(* Logix 5000 project; controller Seperator 1756-L85E rev 33.11; software revision 33.01 *)

TASK IO_Task (periodic, rate 250 ms, priority 2, watchdog 5000 ms) : IO_Simulation
TASK MainTask (continuous, watchdog 5000 ms) : Main_Sequencer, Filler, Capper, Capper_Heads, Filler_Heads1, Filler_Heads2, Filler_Heads3
TASK Process_Control (periodic, rate 250 ms, priority 2, watchdog 5000 ms) : Seperator_Control
TASK RandomTask (event, rate 1 ms, priority 1, watchdog 5000 ms) : RandomProgram   // Random Number Generator
TASK SignalGenerator (periodic, rate 100 ms, priority 1, watchdog 5000 ms) : RandomUpDown
TASK TemperatureLoops (periodic, rate 2000 ms, priority 3, watchdog 5000 ms) : TI101_Temperature

MODULES
   Local : 1756-L85E (ICP 0, rev 33.11)
END_MODULES

TYPE Benchmarks_Comparison :
STRUCT
   Actual_To_Baseline : REAL;
   Actual_To_Same_Interval_Prior_Periods : REAL;
   Production_Lines_To_Like_Lines : REAL;
   Production_Runs_To_Like_Runs : REAL;
END_STRUCT
END_TYPE

TYPE ControllerLEDStatus :
STRUCT
   Off : BOOL;
   SolidGreen : BOOL;
   FlashingGreen : BOOL;
   SolidYellow : BOOL;
   FlashingYellow : BOOL;
   FlashingRed : BOOL;
   SolidRed : BOOL;
END_STRUCT
END_TYPE

TYPE Facility :
STRUCT
   Company_Name : STRING;
   Location_Country : STRING;
   Location_State : STRING;
   Location_City : STRING;
   Benchmarks_Comparison : Benchmarks_Comparison;
   KPIs_Energy_PER_UOP : KPIs_Energy_PER_UOP;
   KPIs_GHG_PER_UOP : KPIs_GHG_PER_UOP;
   WAGES_Demand : WAGES_Demand;
   WAGES_Usage : WAGES_Usage;
END_STRUCT
END_TYPE

TYPE FaultRecord :
STRUCT
   timelow : DINT;
   timehigh : DINT;
   type : INT;
   code : INT;
   info : DINT[8];
END_STRUCT
END_TYPE

TYPE KPIs_Energy_PER_UOP :
STRUCT
   Eunits_PER_UOPunits : REAL;
   Edollar_PER_UOPunits : REAL;
   Eunits_PER_UOPdollar : REAL;
   Edollar_PER_UOPdollar : REAL;
END_STRUCT
END_TYPE

TYPE KPIs_GHG_PER_UOP :
STRUCT
   kG_CO2_e : REAL;
   Metric_Tonnes : REAL;
END_STRUCT
END_TYPE

TYPE Logix_Status_FP :
STRUCT
   ClearMinorFaults : DINT;
   Sts_MinorFaultEvents : DINT;
   Sts_MinorFaultBits : DINT;
   Sts_Redundant : DINT;
   Set_FaceplateAnimation : DINT;
   Val_ProductCode : DINT;
   MemoryTemp : INT[29];
   Val_raw_data : INT;
   Sts_IO_LED_raw : INT;
   Sts_ProductCode : INT;
   Val_Force_data_raw : INT;
   MemoryRequestData : SINT[12];
   Sts_Force_Installed : BOOL;
   Sts_Force_Enabled : BOOL;
   Sts_Faulted : BOOL;
   Sts_Run : BOOL;
   Sts_Program : BOOL;
   Sts_Minor_fault : BOOL;
   Sts_Major_fault : BOOL;
   Sts_KS_in_run : BOOL;
   Sts_KS_in_program : BOOL;
   Sts_KS_in_remote : BOOL;
   Sts_Changingmodes : BOOL;
   Sts_Test : BOOL;
   Sts_Ladder_Working : BOOL;
   Cmd_ClearFaultRecord : BOOL;
   Set_Controller_Description : STRING;
   UpdateDelayTimer : TIMER;
   Val_MajorFault : FaultRecord;
   Val_MFS : FaultRecord;
   Sts_IO_LED : ControllerLEDStatus;
   Sts_Battery_LED : ControllerLEDStatus;
   MemoryData : Memory_Data;
END_STRUCT
END_TYPE

TYPE Memory_Data :
STRUCT
   Free_Mem_IO : DINT;
   Free_Mem_DT : DINT;
   Free_Memory : DINT;
   Total_Mem_IO : DINT;
   Total_Mem_DT : DINT;
   Total_Memory : DINT;
   Biggest_IO_Mem_Size_Ava : DINT;
   Biggest_DT_Mem_Size_Ava : DINT;
END_STRUCT
END_TYPE

TYPE Motor :
STRUCT
   Start : BOOL;
   Stopped : BOOL;
   StartReq : BOOL;
   Alarm : BOOL;
   Running : BOOL;
END_STRUCT
END_TYPE

TYPE Moving_Analog_Indicator :
STRUCT
   Value : REAL;
   Medium_Alarm : REAL;
   High_Alarm : REAL;
   Min : REAL;
   Max : REAL;
END_STRUCT
END_TYPE

TYPE mtrcsdt :
STRUCT
   PartId : STRING;   // Static value per workcell
   IdealCT : REAL;   // Ideal time taken in Seconds to produce each Unit.
   GoodParts : DINT;   // Output Count in Units
   ScrapParts : DINT;   // Reject Count in Units
   TotalParts : DINT;   // Input Count in Units
   Running : BOOL;   // 1=Run Mode
   Monitored_Availability : BOOL;   // 1=Running OR Waiting
   Machine_State : INT;   // [0]=Undefined error [1]=Running [2]=Fault [3]=EfficiencyLoss
   BatchID : STRING;   // Product produced
   Colour : STRING;   // Product colour
   FaultEventTrigger : BOOL;   // 1=Fault detected
   FaultEventValue : INT;   // Fault code
   SlowEventTrigger : BOOL;   // 1=Workcell running slow
   SlowEventValue : INT;   // Slow reason code
   WarningEventTrigger : BOOL;   // 1=Warning detected
   WarningEventValue : INT;   // Warning code
END_STRUCT
END_TYPE

TYPE Phase_Control :
STRUCT
   Cmd_Start : BOOL;
   Cmd_Stop : BOOL;
   Cmd_Reset : BOOL;
END_STRUCT
END_TYPE

TYPE STRING_12 :
STRUCT
   LEN : DINT;
   DATA : SINT[12];
END_STRUCT
END_TYPE

TYPE STRING_16_UDT :
STRUCT
   LEN : DINT;
   DATA : SINT[16];
END_STRUCT
END_TYPE

TYPE STRING_20 :
STRUCT
   LEN : DINT;
   DATA : SINT[20];
END_STRUCT
END_TYPE

TYPE STRING_40 :
STRUCT
   LEN : DINT;
   DATA : SINT[40];
END_STRUCT
END_TYPE

TYPE Valve :
STRUCT
   Open : BOOL;
   Closed : BOOL;
   OpenReq : BOOL;
   Alarm : BOOL;
   Opened : BOOL;
END_STRUCT
END_TYPE

TYPE WAGES_Demand :
STRUCT
   Water_Demand : REAL;
   Air_Demand : REAL;
   Gas_Demand : REAL;
   Electric_Demand : REAL;
   Steam_Demand : REAL;
END_STRUCT
END_TYPE

TYPE WAGES_Usage :
STRUCT
   Water_Usage : REAL;
   Air_Usage : REAL;
   Gas_Usage : REAL;
   Electric_Usage : REAL;
   Steam_Usage : REAL;
END_STRUCT
END_TYPE

ADD_ON_INSTRUCTION AOI_SIM_RNG_Simple   (* revision 1.3, vendor Dr. Frank Jordan / Rockwell Automation, ExecutePrescan *)
// Simple Random Number Generator
// Revision note:
// This code is provided as application example without any warranty
// Help:
// George Marsaglia 's MWC (multiply with carry) algorithm
// (taken from http://www.codeproject.com/Articles/25172/Simple-Random-Number-Generation)
VAR_INPUT
   Seed : ALIAS FOR LocalSeed; {access Read Only, visible}
END_VAR
VAR_OUTPUT
   Count : DINT; {access Read Only, visible}
   Number : REAL; {access Read Only, visible}
END_VAR
VAR_INPUT
   TriggerSeed : ALIAS FOR LocalTriggerSeed; {access Read Only, visible}
   Reset : ALIAS FOR LocalReset; {access Read Only, visible}
END_VAR
VAR
   m_z : DINT; {access None}
   m_w : DINT; {access None}
   delta : REAL; {access None}
   consB : DINT; {access None}
   consA : DINT; {access None}
   AOI_UMUL : UMUL; {access None}
   u : DINT; {access None}
   AOI_UADD : UADD; {access None}
   LocalTriggerSeed : BOOL; {access Read Only}
   LocalSeed : DINT; {access Read Only}
   LocalReset : BOOL; {access Read Only}
   tmp : DINT; {access None}
   Overflow : BOOL; {access None}
END_VAR

ROUTINE Logic   (* ladder *)
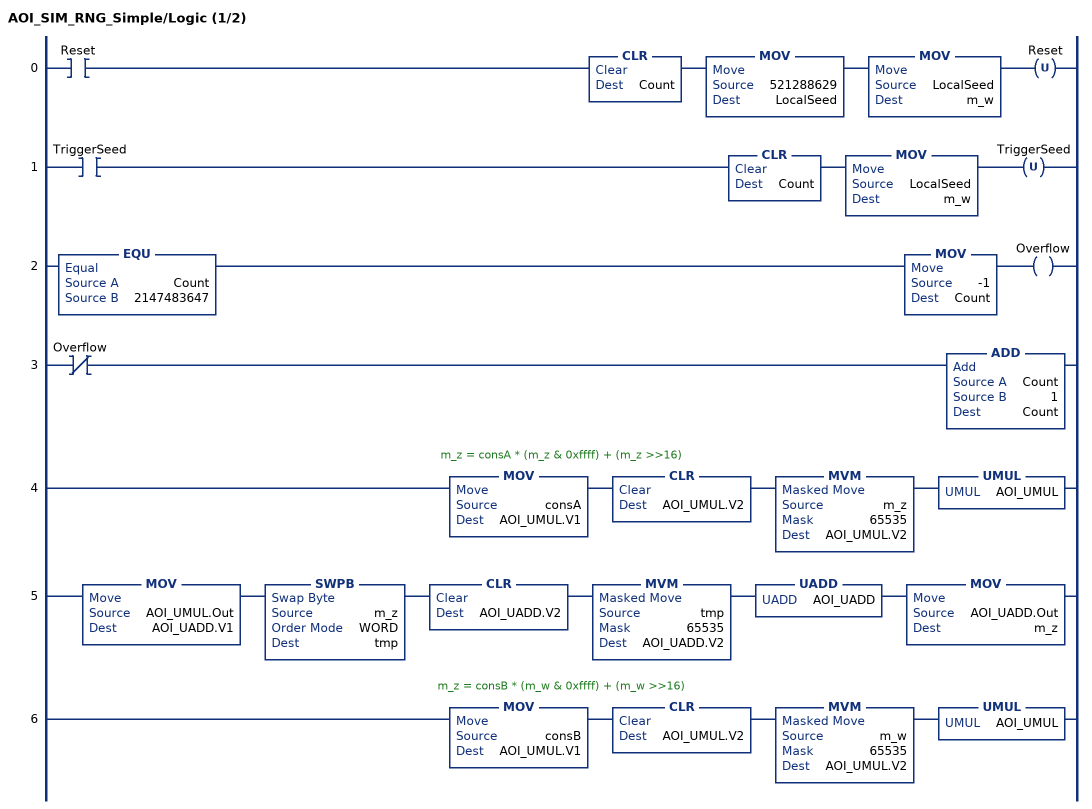
   0: XIC(Reset)CLR(Count)MOV(521288629,LocalSeed)MOV(LocalSeed,m_w)OTU(Reset);
   1: XIC(TriggerSeed)CLR(Count)MOV(LocalSeed,m_w)OTU(TriggerSeed);
   2: EQU(Count,2147483647)MOV(-1,Count)OTE(Overflow);
   3: XIO(Overflow)ADD(Count,1,Count);
   // m_z = consA * (m_z & 0xffff) + (m_z >>16)
   4: MOV(consA,AOI_UMUL.V1)CLR(AOI_UMUL.V2)MVM(m_z,65535,AOI_UMUL.V2)UMUL(AOI_UMUL);
   5: MOV(AOI_UMUL.Out,AOI_UADD.V1)SWPB(m_z,WORD,tmp)CLR(AOI_UADD.V2)MVM(tmp,65535,AOI_UADD.V2)UADD(AOI_UADD)MOV(AOI_UADD.Out,m_z);
   // m_z = consB * (m_w & 0xffff) + (m_w >>16)
   6: MOV(consB,AOI_UMUL.V1)CLR(AOI_UMUL.V2)MVM(m_w,65535,AOI_UMUL.V2)UMUL(AOI_UMUL);
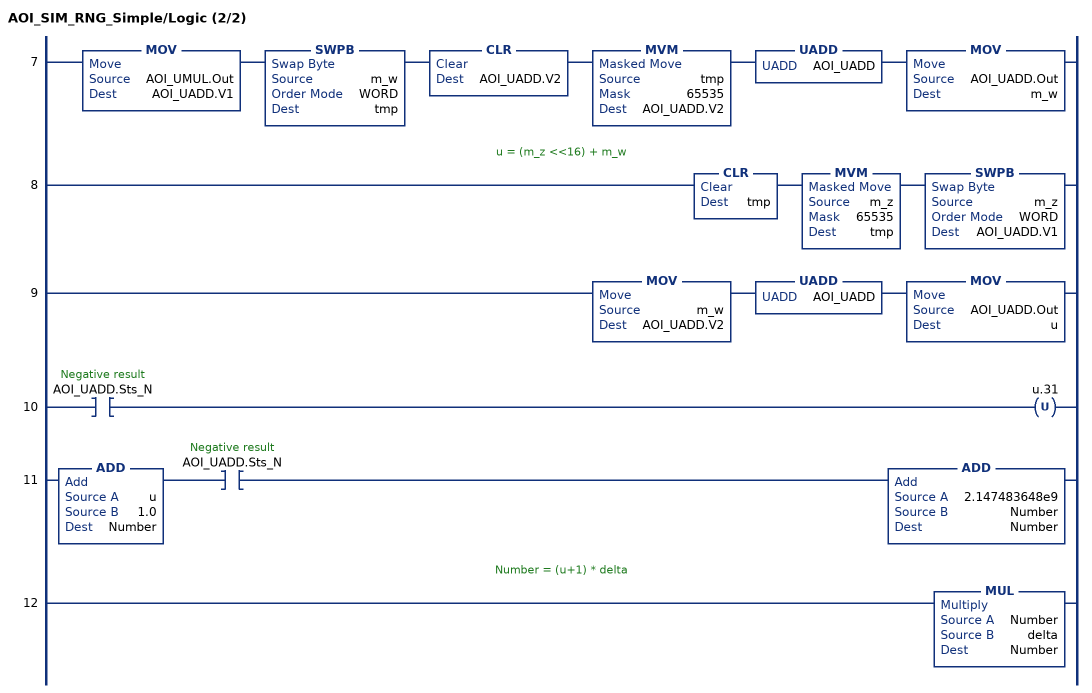
   7: MOV(AOI_UMUL.Out,AOI_UADD.V1)SWPB(m_w,WORD,tmp)CLR(AOI_UADD.V2)MVM(tmp,65535,AOI_UADD.V2)UADD(AOI_UADD)MOV(AOI_UADD.Out,m_w);
   // u = (m_z <<16) + m_w
   8: CLR(tmp)MVM(m_z,65535,tmp)SWPB(m_z,WORD,AOI_UADD.V1);
   9: MOV(m_w,AOI_UADD.V2)UADD(AOI_UADD)MOV(AOI_UADD.Out,u);
   10: XIC(AOI_UADD.Sts_N)OTU(u.31);
   11: ADD(u,1.0,Number)XIC(AOI_UADD.Sts_N)ADD(2.147483648e9,Number,Number);
   // Number = (u+1) * delta
   12: MUL(Number,delta,Number);
END_ROUTINE

ROUTINE Prescan   (* ladder *)
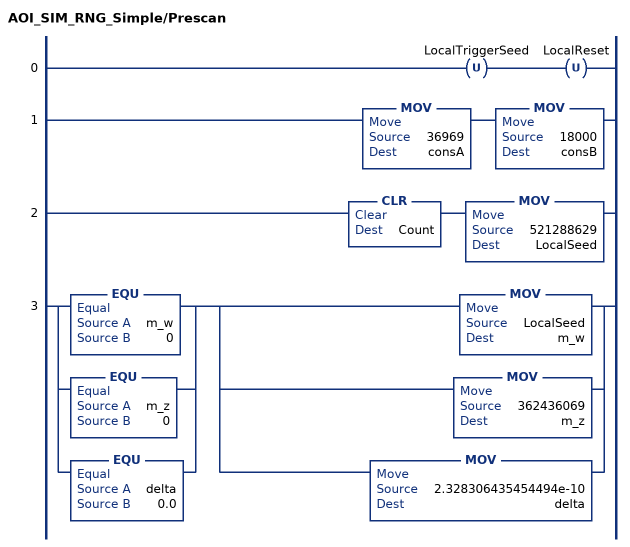
   0: OTU(LocalTriggerSeed)OTU(LocalReset);
   1: MOV(36969,consA)MOV(18000,consB);
   2: CLR(Count)MOV(521288629,LocalSeed);
   3: [EQU(m_w,0) ,EQU(m_z,0) ,EQU(delta,0.0) ][MOV(LocalSeed,m_w) ,MOV(362436069,m_z) ,MOV(2.328306435454494e-10,delta) ];
END_ROUTINE
END_ADD_ON_INSTRUCTION

ADD_ON_INSTRUCTION FTV_ctrl   (* revision 1.0 *)
VAR_INPUT
   nr_of_screens : DINT := 1; {visible}
   ActiveScreen : DINT;
   ScreenOverride : DINT;
   delay : DINT := 10; {visible}
   ScreenRequest : DINT;
END_VAR
VAR_OUTPUT
   Act : BOOL; {visible}
END_VAR
VAR
   Screen_delay : FBD_TIMER; {access None}
END_VAR

ROUTINE Logic   (* structured text *)
   Act:= (ActiveScreen >=100);
   
   Screen_delay.PRE:=delay*1000;
   Screen_delay.TimerEnable:=Act & NOT Screen_delay.DN & (ScreenRequest=0);
   TONR(Screen_delay);
   IF Act AND ScreenOverride<100 THEN ScreenOverride:=100;END_IF;
   IF Screen_delay.DN THEN ScreenOverride:= ScreenOverride+1;END_IF;
   IF ScreenOverride>=(100+ nr_of_screens) THEN ScreenOverride:=100;END_IF;
   
   IF ScreenRequest <> 0 THEN ScreenOverride:=ScreenRequest;
   	IF ActiveScreen=ScreenRequest THEN
   		ScreenOverride:=0;
   		ScreenRequest:=0;
   	END_IF;
   END_IF;
   
   IF NOT Act THEN ScreenOverride:=0; END_IF;
END_ROUTINE
END_ADD_ON_INSTRUCTION

ADD_ON_INSTRUCTION MotorSim   (* revision 1.0, vendor Rockwell, ExecutePrescan *)
VAR_INPUT
   MotorStartRequest : BOOL; {visible}
END_VAR
VAR_OUTPUT
   MotorRunning : BOOL; {access Read Only, visible}
   MotorStopped : BOOL; {access Read Only, visible}
END_VAR
VAR
   StartCommand : BOOL;
   RunningCommandDelay : TIMER := (PRE := 2000);
   StoppedCommandDelay : TIMER := (PRE := 2000);
END_VAR

ROUTINE Logic   (* ladder *)
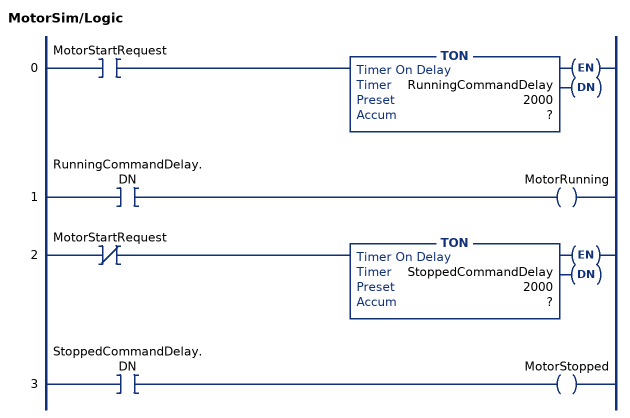
   0: XIC(MotorStartRequest)TON(RunningCommandDelay,?,?);
   1: XIC(RunningCommandDelay.DN)OTE(MotorRunning);
   2: XIO(MotorStartRequest)TON(StoppedCommandDelay,?,?);
   3: XIC(StoppedCommandDelay.DN)OTE(MotorStopped);
END_ROUTINE

ROUTINE Prescan   (* structured text *)
   RunningCommandDelay.PRE:=2000;
   StoppedCommandDelay.PRE:=2000;
   
END_ROUTINE
END_ADD_ON_INSTRUCTION

ADD_ON_INSTRUCTION P_Alarm   (* revision 3.0 02 Release, vendor Rockwell Automation, ExecutePrescan, ExecuteEnableInFalse *)
// Alarm
// Revision note:
// Changed suppress to shelve, inhibit to suppress (ISA 18.2-2009 and FTView 7 alignment), added auto unshelve timer, program command to unshelve. Removed: Ack on shelve. Added: clear Alm when disabled, PCfg_AllowExist, Cfg_Tag, Cfg_Cond, Inf_Lib, Inf_Type. Added Com_AE Local Tag for FTAE communication. Changed Cfg_MaxShelfT check to LEQ 0.  (INT 1 to 32767 is valid.)
// Help:
// Copyright © Rockwell Automation, Inc.  All Rights Reserved.
// This instruction monitors one input condition and provides one Alarm with:
//   * configurable latching (reset required) and acknowledgement requirement
//   * configurable alarm severity
//       1 = Low  (blue, typ. informational)
//       2 = Medium  (yelllow, typ. warning)
//       3 = High  (red, typ. process exception)
//       4 = Highest  (magenta, typ. equip. fault)
//   * configurable minimum ON time (e.g., to ensure it is seen by the HMI)
//   * commands to suppress/unsuppress (Prog), shelve/unshelve (Oper)
//         and disable/enable (Maint) the alarm.
//   * configurable amount of time shelved to automatically unshelve an alarm
//   * FTA&E support for suppressed, shelved and disabled states (V7.0)
// NOTE regarding parameter naming:
//   FTAE names (same as ALMD instruction) are used instead
//   of the ANSI/ISA 18.2-2009 names, as follows:
//    "Disabled" is the equivalent of "Out of Service" in ISA 18.2.
//       (The Disabled state is owned by Maintenance.)
//    "Suppressed" is the equivalent of "Suppressed by Design" in
//       ISA 18.2. (The Suppressed state is owned by Program logic.)
//    "Shelved" is the same as in ISA 18.2.
//       (The Shelved state is owned by Operator, but may be cleared
//       by Program logic based on time, shift change, etc.)
// This instruction is usually nested within other instructions, with one instance
// used for each Alarm generated by the containing instruction.  It may also be
// used as a standalone instruction for Alarm conditions generated by custom logic.
// FTAE Alarm Setup:
//   (object).(alarm).Com_AE.0:  Alarm to FTAE
//     .Com_AE.1:   Ack to/from FTAE
//     .Com_AE.3:   Shelved from FTAE Status
//     .Com_AE.4:   Shelve/Reshelve to FTAE Control (auto reset)
//     .Com_AE.5:   Unshelve to FTAE Control (auto reset)
//     .Com_AE.6:   Suppressed to/from FTAE
//     .Com_AE.8:   Unsuppress to FTAE Control (auto reset)
//     .Com_AE.9:   Disabled to/from FTAE
//     .Com_AE.11: Enable to FTAE Control (auto reset)
//    all other bits unused
//     .Cfg_MaxShelfT is also used in FTAE config.
VAR_INPUT
   Inp : BOOL := 1; {visible}   // Alarm Condition Input 1=Alarm
   Inp_Reset : BOOL; {visible}   // 1=Reset Alarm requiring reset
   Cfg_Exists : BOOL := 1;   // 1=Alarm configured to exist, 0=Does not exist, don't scan
   Cfg_ResetReqd : BOOL;   // 1=Latched Alarm, a Reset is required to clear this Alarm
   Cfg_AckReqd : BOOL := 1;   // 1=Acknowledge required for this Alarm
   Cfg_AllowShelve : BOOL := 1;   // 1=Allow Operator to Shelve this Alarm
   Cfg_AllowDisable : BOOL := 1;   // 1=Allow Maintenance to Disable this Alarm
   Cfg_PCmdClear : BOOL := 1;   // 1=Clear Program Commands on receipt 0=Leave Set
   Cfg_Severity : SINT := 3;   // Alarm Severity: 1=Low, 2=Medium, 3=High, 4=Highest
   Cfg_AlmMinOnT : DINT := 5;   // Minimum time Alm output stays on (sec)
   Cfg_MaxShelfT : INT := 480;   // Auto unshelve after shelved this long (1..32767 minutes)
   PCfg_AllowExist : BOOL := 1;   // 1=Alarm can be configured to exist, 0=other configs make alarm meaningless
   PCmd_Reset : BOOL;   // Program Command to Reset latched alarm
   PCmd_Ack : BOOL;   // Program Command to Acknowledge alarm
   PCmd_Suppress : BOOL;   // Program Command to Suppress by Design (inhibits new alarm)
   PCmd_Unsuppress : BOOL;   // Program Command to Unsuppress (allows new alarm)
   PCmd_Unshelve : BOOL;   // Program Command to Unshelve (e.g., on shift change)
   OCmd_Reset : BOOL;   // Operator Command to Reset latched alarm
   OCmd_Ack : BOOL;   // Operator Command to Acknowledge alarm
   OCmd_Shelve : BOOL;   // Operator Command to Shelve Alarm (inhibits new alarm)
   OCmd_Unshelve : BOOL;   // Operator Command to Unshelve alarm (allows new alarm)
   MCmd_Disable : BOOL;   // Maintenance Command to Disable alarm (inhibits new alarm)
   MCmd_Enable : BOOL;   // Maintenance Command to Enable alarm (allows new alarm)
END_VAR
VAR_OUTPUT
   Val_Notify : SINT; {access Read Only}   // Current Alarm Severity and Acknowledgement (enumeration)
   Val_MinToUnshelve : DINT; {access Read Only, visible}   // Number of minutes until this alarm unshelves itself (mmm:ss)
   Val_SecToUnshelve : DINT; {access Read Only, visible}   // Number of Seconds until this alarm unshelves itself (mmm:ss)
   Alm : ALIAS FOR Com_AE.0; {visible}   // Alarm output 1=In Alarm
   Ack : ALIAS FOR Com_AE.1; {visible}   // Alarm acknowledged status: 1=Ack rcvd
   Shelved : ALIAS FOR Com_AE.3; {visible}   // 1=Alarm has been Shelved by Operator (inhibits new alarm)
   Suppressed : ALIAS FOR Com_AE.6; {visible}   // 1=Alarm has been Suppressed by Program (inhibits new alarm)
   Disabled : ALIAS FOR Com_AE.9; {visible}   // 1=Alarm has been Disabled by Maintanance (inhibits new alarm)
   Sts_AlmInh : BOOL; {access Read Only}   // 1=Alarm has been suppressed, shelved or disabled, display "I" icon
   Sts_Err : BOOL; {access Read Only}   // 1=Error in Config: see detail Err_ bits for reason
   Err_Timer : BOOL; {access Read Only}   // 1=Error in Config: Alarm Min On Time, Shelf Time (use 0 to 2147483)
   Err_Severity : BOOL; {access Read Only}   // 1=Error in Config: Invalid Severity (use 1 to 4)
   Rdy_Reset : BOOL; {access Read Only}   // Ready to receive OCmd_Reset (enables button)
   Rdy_Ack : BOOL; {access Read Only}   // Ready to receive OCmd_Ack (enables button)
   Rdy_Shelve : BOOL; {access Read Only}   // Ready to receive OCmd_Shelve (enables button)
   Rdy_Unshelve : BOOL; {access Read Only}   // Ready to receive OCmd_Unshelve (enables button)
   Rdy_Disable : BOOL; {access Read Only}   // Ready to receive MCmd_Disable (enables button)
   Rdy_Enable : BOOL; {access Read Only}   // Ready to receive MCmd_Enable (enables button)
   P_Alarm : BOOL;   // Unique Parameter Name for auto - discovery
END_VAR
VAR
   Wrk_Alm : BOOL; {access None}   // Internal Alarm Status
   Wrk_Suppressed : BOOL; {access None}   // Internal Alarm Suppressed Status
   Wrk_AlmMinOnT : TIMER := (PRE := 5000); {access None}   // Alarm output minimum ON time to be seen by alarm server
   Wrk_AutoAckT : TIMER := (PRE := 5000); {access None}   // Time to clear Ack bit when Ack not required
   Wrk_ShelfT : TIMER; {access None}   // Time to auto Unshelve a Shelved Alarm
   Inf_Tab : SINT;   // Tab to display (FTView ME)
   Com_AE : INT := 2#0000_0000_0000_0010;   // Communication with HMI / Alarm/Event Server (see bit descriptions)
        .10   // (not used)
        .11   // Enable to AE Control
        .12   // (not used)
        .13   // (not used)
        .14   // (not used)
        .15   // (not used)
        .0   // Alarm to AE
        .1   // Acked from AE Status, Ack to AE Control
        .2   // (not used)
        .3   // Shelved from AE Status
        .4   // Shelve to AE Control
        .5   // Unshelve to AE Control
        .6   // Suppressed from AE Status, Suppress to AE Control
        .7   // (not used)
        .8   // Unsuppress to AE Control
        .9   // Disabled from AE Status, Disable to AE Control
   Cfg_Tag : STRING_20 := 'P_Alarm';   // Alarm Tag Text (e.g., "LAHH-101")
   Cfg_Cond : STRING_20 := 'Alarm Condition';   // Alarm Condition Text (e.g., "High-High PV")
   Wrk_SecToUnshelve : DINT; {access None}   // Number of seconds until this alarm unshelves itself
   Inf_Lib : STRING_12 := 'RA-BAS'; {access Read Only}   // Display Library for Faceplate call-up
   Inf_Type : STRING_16_UDT := 'P_Alarm'; {access Read Only}   // Must contain AOI name, used for HMI and Information S/W
END_VAR

ROUTINE EnableInFalse   (* ladder *)
// Perform Alarm processing, but Invert Alarm Input ("Inp") for use on LD rung (EnableIn False)
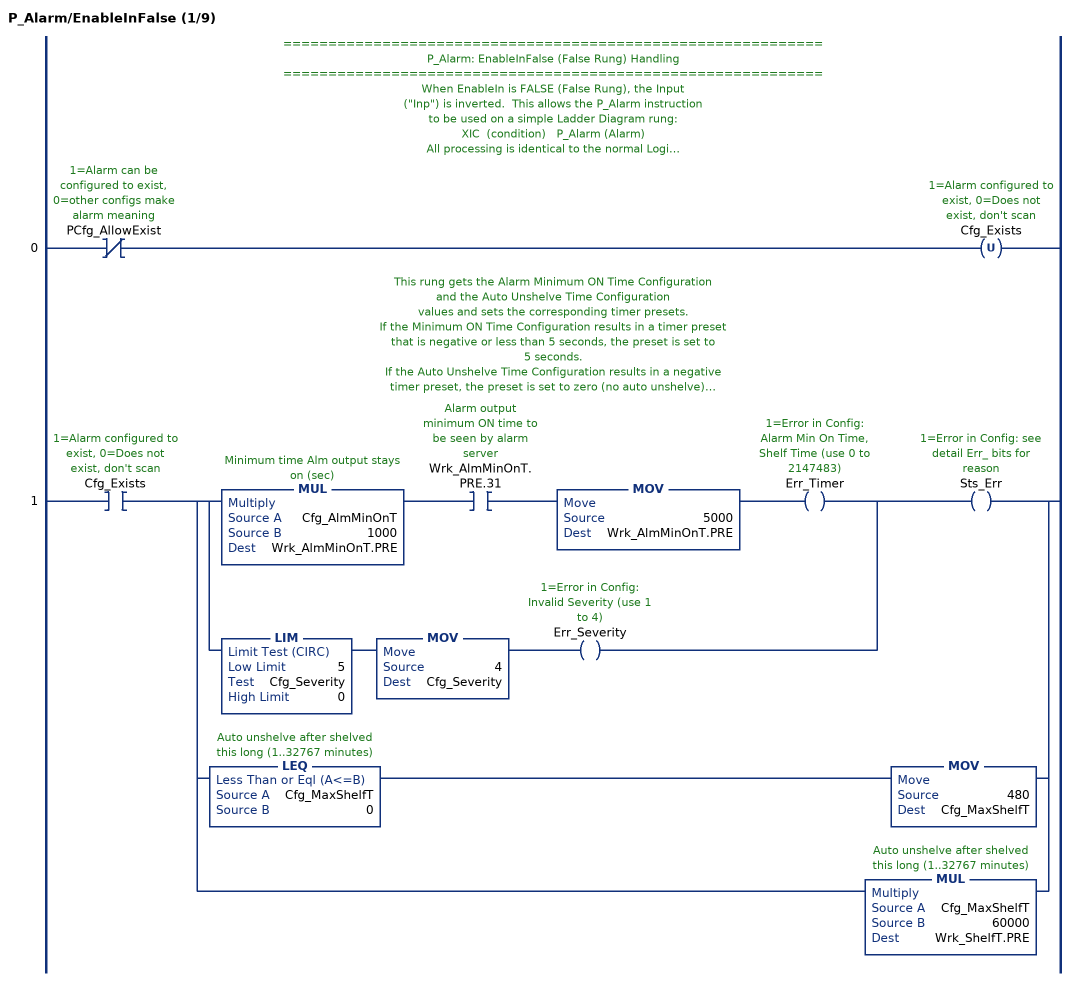
   // ============================================================
   // P_Alarm: EnableInFalse (False Rung) Handling
   // ============================================================
   // When EnableIn is FALSE (False Rung), the Input
   // ("Inp") is inverted.  This allows the P_Alarm instruction
   // to be used on a simple Ladder Diagram rung:
   // XIC  (condition)   P_Alarm (Alarm)
   // All processing is identical to the normal Logic
   // routine, except references to Inp are inverted!
   // ============================================================
   // CONFIGURATION
   // ============================================================
   // In the object containing this alarm, other configuration (such as not having
   // any limit switches) may make this particular alarm meaningless.
   // The Program Configuration "Allow Exist" is used to hide this alarm
   // on the object's faceplate and other graphics, and forces the Cfg_Exist to 0.
   // #####  V3.0-00  2013-06-30:  Added PCfg_AllowExist.  #####
   0: XIO(PCfg_AllowExist)OTU(Cfg_Exists);
   // This rung gets the Alarm Minimum ON Time Configuration
   // and the Auto Unshelve Time Configuration
   // values and sets the corresponding timer presets.
   // If the Minimum ON Time Configuration results in a timer preset
   // that is negative or less than 5 seconds, the preset is set to
   // 5 seconds.
   // If the Auto Unshelve Time Configuration results in a negative
   // timer preset, the preset is set to zero (no auto unshelve).
   //   The bad Config is flagged (Err_Timer).
   // Bad Config is also flagged if the Cfg_Severity is out of range (valid = 1..4)
   // #####  V3.0-00  2013-06-30:  Changed Program Inhibit to Suppress, Operator Suppress to Shelve.  #####
   // #####  Added Shelf Timer config check; if Severity out of range, make it "Fault".  #####
   // #####  V3.0-02  2013-10-30:  Changed Cfg_MaxShelfT check to LEQ 0.  (INT 1 to 32767 is valid.)  #####
   1: XIC(Cfg_Exists)[[MUL(Cfg_AlmMinOnT,1000,Wrk_AlmMinOnT.PRE) XIC(Wrk_AlmMinOnT.PRE.31) MOV(5000,Wrk_AlmMinOnT.PRE) OTE(Err_Timer) ,LIM(5,Cfg_Severity,0) MOV(4,Cfg_Severity) OTE(Err_Severity) ] OTE(Sts_Err) ,LEQ(Cfg_MaxShelfT,0) MOV(480,Cfg_MaxShelfT) ,MUL(Cfg_MaxShelfT,60000,Wrk_ShelfT.PRE) ];
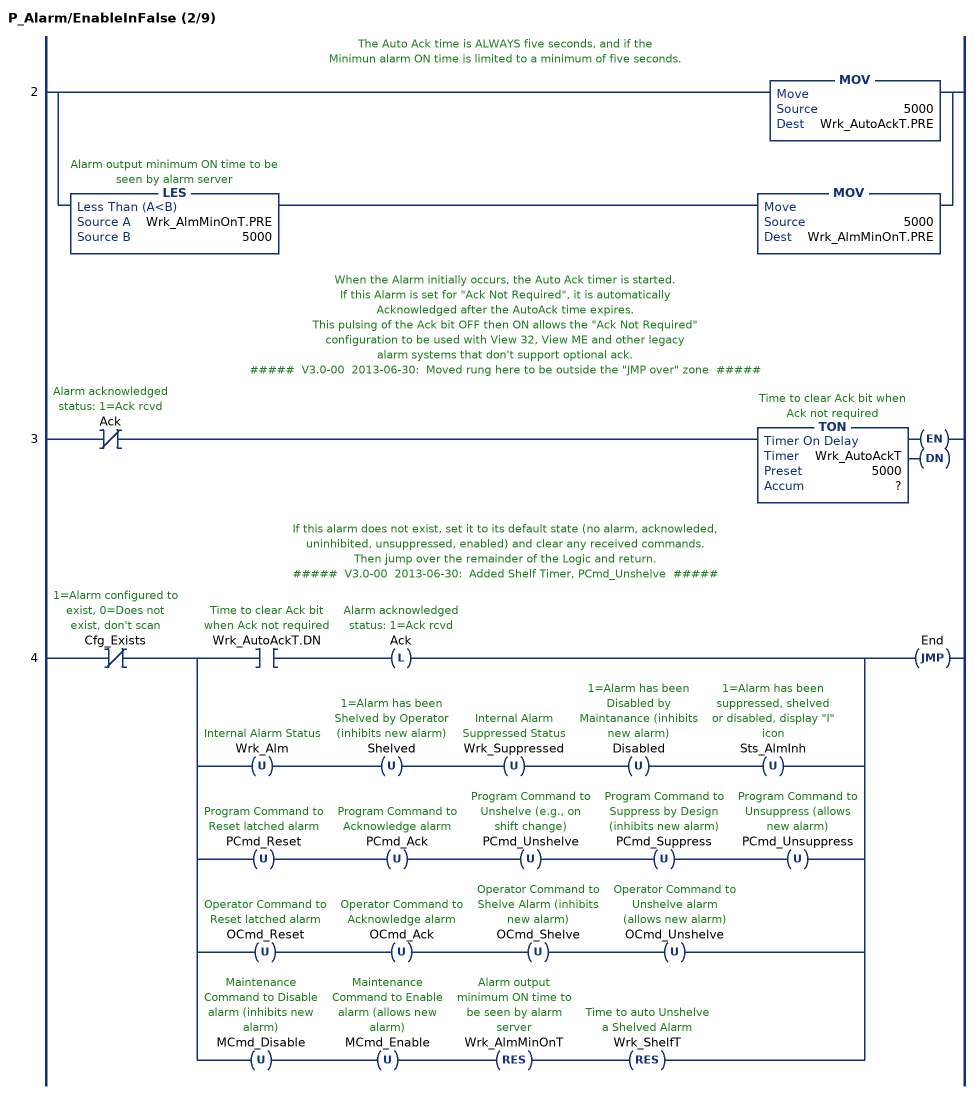
   // The Auto Ack time is ALWAYS five seconds, and if the
   // Minimun alarm ON time is limited to a minimum of five seconds.
   2: [MOV(5000,Wrk_AutoAckT.PRE) ,LES(Wrk_AlmMinOnT.PRE,5000) MOV(5000,Wrk_AlmMinOnT.PRE) ];
   // When the Alarm initially occurs, the Auto Ack timer is started.
   // If this Alarm is set for "Ack Not Required", it is automatically
   // Acknowledged after the AutoAck time expires.
   // This pulsing of the Ack bit OFF then ON allows the "Ack Not Required"
   // configuration to be used with View 32, View ME and other legacy
   // alarm systems that don't support optional ack.
   // #####  V3.0-00  2013-06-30:  Moved rung here to be outside the "JMP over" zone  #####
   3: XIO(Ack)TON(Wrk_AutoAckT,?,?);
   // If this alarm does not exist, set it to its default state (no alarm, acknowleded,
   // uninhibited, unsuppressed, enabled) and clear any received commands.
   // Then jump over the remainder of the Logic and return.
   // #####  V3.0-00  2013-06-30:  Added Shelf Timer, PCmd_Unshelve  #####
   4: XIO(Cfg_Exists)[XIC(Wrk_AutoAckT.DN) OTL(Ack) ,OTU(Wrk_Alm) OTU(Shelved) OTU(Wrk_Suppressed) OTU(Disabled) OTU(Sts_AlmInh) ,OTU(PCmd_Reset) OTU(PCmd_Ack) OTU(PCmd_Unshelve) OTU(PCmd_Suppress) OTU(PCmd_Unsuppress) ,OTU(OCmd_Reset) OTU(OCmd_Ack) OTU(OCmd_Shelve) OTU(OCmd_Unshelve) ,OTU(MCmd_Disable) OTU(MCmd_Enable) RES(Wrk_AlmMinOnT) RES(Wrk_ShelfT) ]JMP(End);
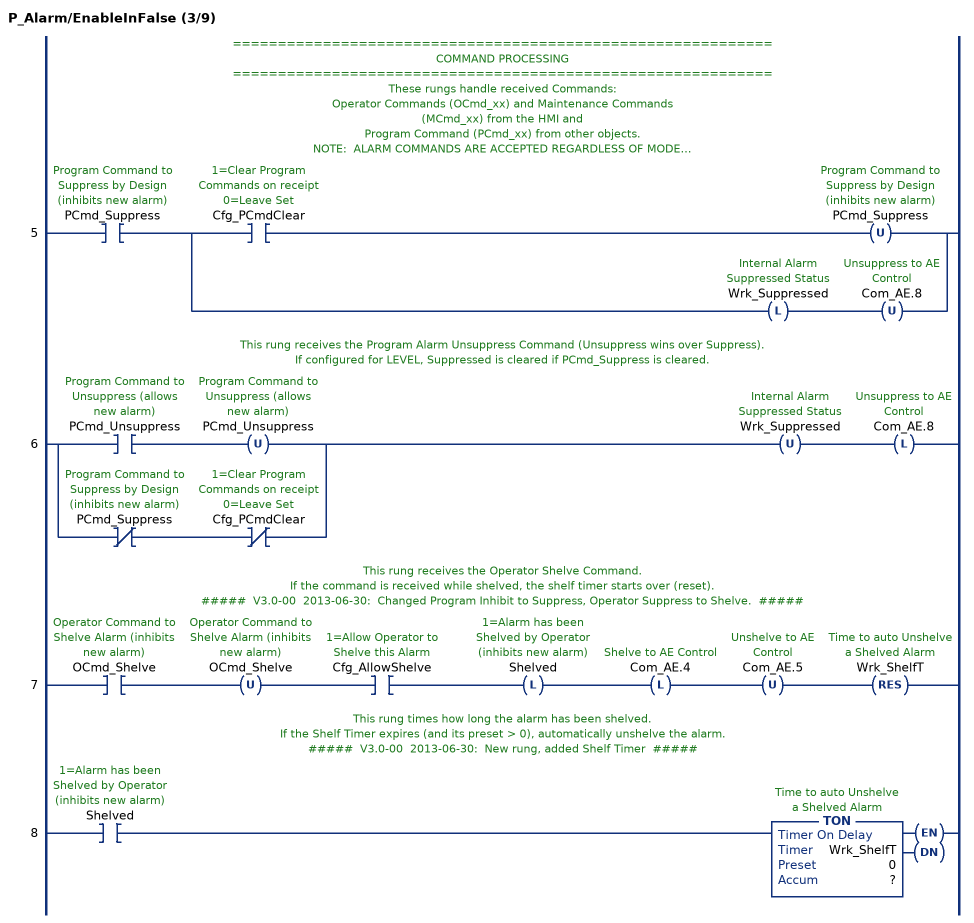
   // ============================================================
   // COMMAND PROCESSING
   // ============================================================
   // These rungs handle received Commands:
   // Operator Commands (OCmd_xx) and Maintenance Commands
   // (MCmd_xx) from the HMI and
   // Program Command (PCmd_xx) from other objects.
   // NOTE:  ALARM COMMANDS ARE ACCEPTED REGARDLESS OF MODE.
   // This rung receives the Program Alarm Inhibit Command.
   // If configured for EDGE, the Command is cleared.
   5: XIC(PCmd_Suppress)[XIC(Cfg_PCmdClear) OTU(PCmd_Suppress) ,OTL(Wrk_Suppressed) OTU(Com_AE.8) ];
   // This rung receives the Program Alarm Unsuppress Command (Unsuppress wins over Suppress).
   // If configured for LEVEL, Suppressed is cleared if PCmd_Suppress is cleared.
   6: [XIC(PCmd_Unsuppress) OTU(PCmd_Unsuppress) ,XIO(PCmd_Suppress) XIO(Cfg_PCmdClear) ]OTU(Wrk_Suppressed)OTL(Com_AE.8);
   // This rung receives the Operator Shelve Command.
   // If the command is received while shelved, the shelf timer starts over (reset).
   // #####  V3.0-00  2013-06-30:  Changed Program Inhibit to Suppress, Operator Suppress to Shelve.  #####
   7: XIC(OCmd_Shelve)OTU(OCmd_Shelve)XIC(Cfg_AllowShelve)OTL(Shelved)OTL(Com_AE.4)OTU(Com_AE.5)RES(Wrk_ShelfT);
   // This rung times how long the alarm has been shelved.
   // If the Shelf Timer expires (and its preset > 0), automatically unshelve the alarm.
   // #####  V3.0-00  2013-06-30:  New rung, added Shelf Timer  #####
   8: XIC(Shelved)TON(Wrk_ShelfT,?,?);
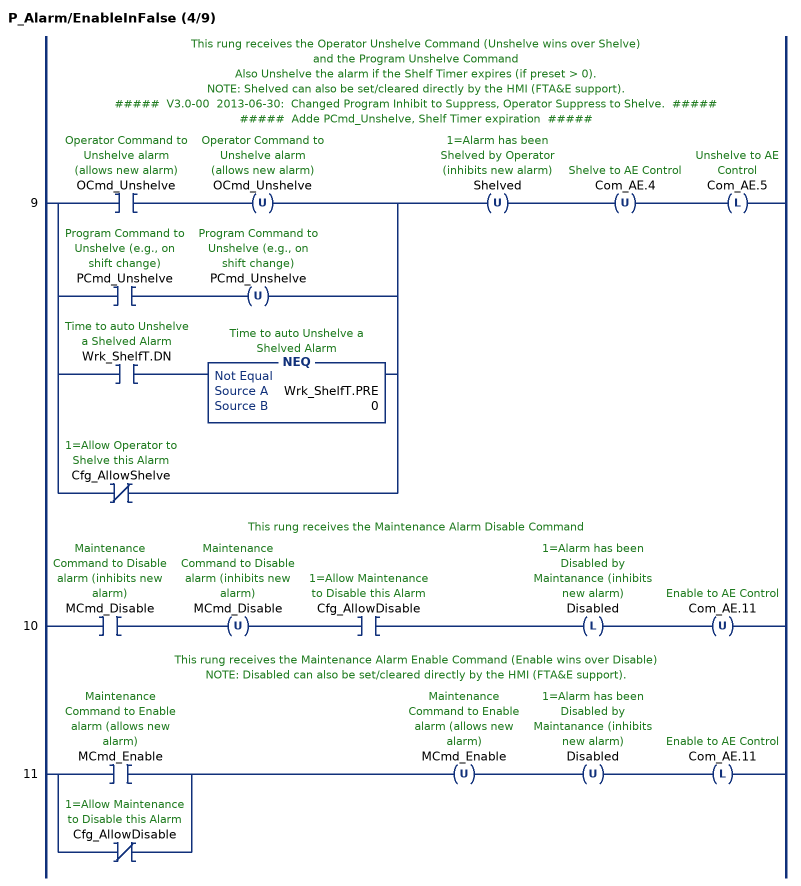
   // This rung receives the Operator Unshelve Command (Unshelve wins over Shelve)
   // and the Program Unshelve Command
   // Also Unshelve the alarm if the Shelf Timer expires (if preset > 0).
   // NOTE: Shelved can also be set/cleared directly by the HMI (FTA&E support).
   // #####  V3.0-00  2013-06-30:  Changed Program Inhibit to Suppress, Operator Suppress to Shelve.  #####
   // #####  Adde PCmd_Unshelve, Shelf Timer expiration  #####
   9: [XIC(OCmd_Unshelve) OTU(OCmd_Unshelve) ,XIC(PCmd_Unshelve) OTU(PCmd_Unshelve) ,XIC(Wrk_ShelfT.DN) NEQ(Wrk_ShelfT.PRE,0) ,XIO(Cfg_AllowShelve) ]OTU(Shelved)OTU(Com_AE.4)OTL(Com_AE.5);
   // This rung receives the Maintenance Alarm Disable Command
   10: XIC(MCmd_Disable)OTU(MCmd_Disable)XIC(Cfg_AllowDisable)OTL(Disabled)OTU(Com_AE.11);
   // This rung receives the Maintenance Alarm Enable Command (Enable wins over Disable)
   // NOTE: Disabled can also be set/cleared directly by the HMI (FTA&E support).
   11: [XIC(MCmd_Enable) ,XIO(Cfg_AllowDisable) ]OTU(MCmd_Enable)OTU(Disabled)OTL(Com_AE.11);
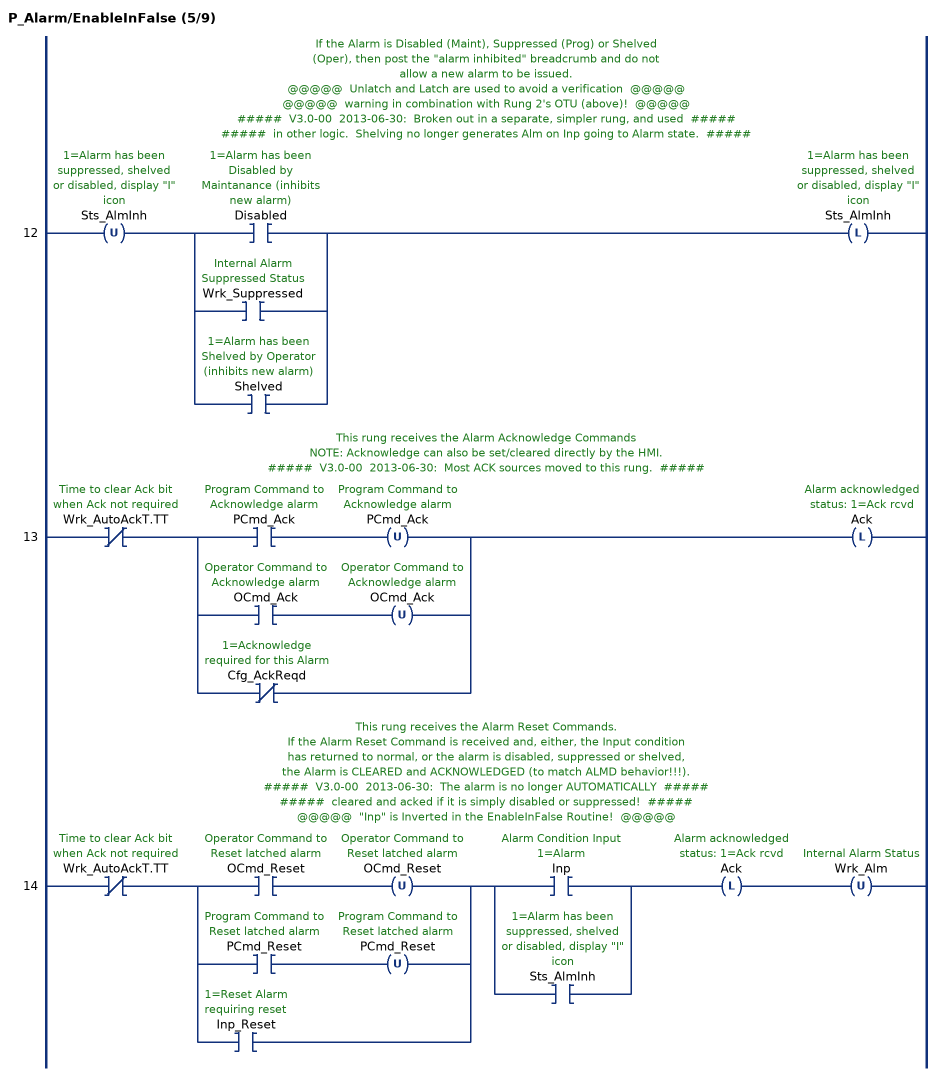
   // If the Alarm is Disabled (Maint), Suppressed (Prog) or Shelved
   // (Oper), then post the "alarm inhibited" breadcrumb and do not
   // allow a new alarm to be issued.
   // @@@@@  Unlatch and Latch are used to avoid a verification  @@@@@
   // @@@@@  warning in combination with Rung 2's OTU (above)!  @@@@@
   // #####  V3.0-00  2013-06-30:  Broken out in a separate, simpler rung, and used  #####
   // #####  in other logic.  Shelving no longer generates Alm on Inp going to Alarm state.  #####
   12: OTU(Sts_AlmInh)[XIC(Disabled) ,XIC(Wrk_Suppressed) ,XIC(Shelved) ]OTL(Sts_AlmInh);
   // This rung receives the Alarm Acknowledge Commands
   // NOTE: Acknowledge can also be set/cleared directly by the HMI.
   // #####  V3.0-00  2013-06-30:  Most ACK sources moved to this rung.  #####
   13: XIO(Wrk_AutoAckT.TT)[XIC(PCmd_Ack) OTU(PCmd_Ack) ,XIC(OCmd_Ack) OTU(OCmd_Ack) ,XIO(Cfg_AckReqd) ]OTL(Ack);
   // This rung receives the Alarm Reset Commands.
   // If the Alarm Reset Command is received and, either, the Input condition
   // has returned to normal, or the alarm is disabled, suppressed or shelved,
   // the Alarm is CLEARED and ACKNOWLEDGED (to match ALMD behavior!!!).
   // #####  V3.0-00  2013-06-30:  The alarm is no longer AUTOMATICALLY  #####
   // #####  cleared and acked if it is simply disabled or suppressed!  #####
   // @@@@@  "Inp" is Inverted in the EnableInFalse Routine!  @@@@@
   14: XIO(Wrk_AutoAckT.TT)[XIC(OCmd_Reset) OTU(OCmd_Reset) ,XIC(PCmd_Reset) OTU(PCmd_Reset) ,XIC(Inp_Reset) ][XIC(Inp) ,XIC(Sts_AlmInh) ]OTL(Ack)OTU(Wrk_Alm);
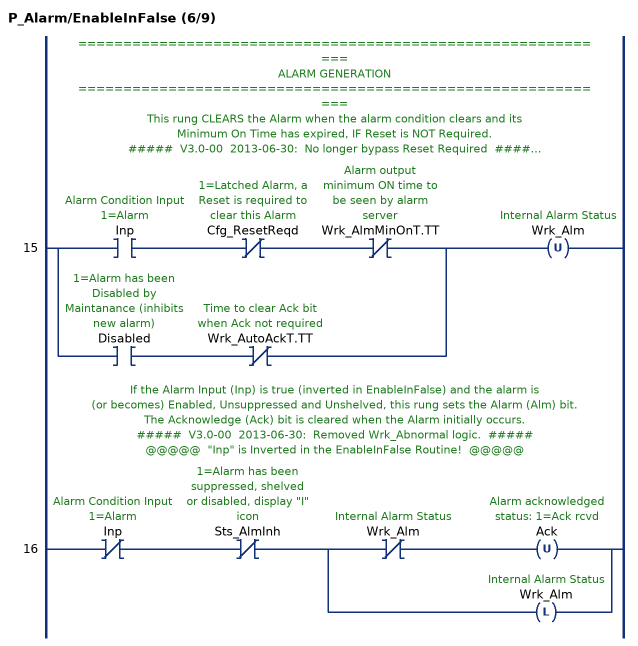
   // ============================================================
   // ALARM GENERATION
   // ============================================================
   // This rung CLEARS the Alarm when the alarm condition clears and its
   // Minimum On Time has expired, IF Reset is NOT Required.
   // #####  V3.0-00  2013-06-30:  No longer bypass Reset Required  #####
   // #####  when the alarm is Shelved by the Operator.  #####
   // @@@@@  "Inp" is Inverted in the EnableInFalse Routine!  @@@@@
   15: [XIC(Inp) XIO(Cfg_ResetReqd) XIO(Wrk_AlmMinOnT.TT) ,XIC(Disabled) XIO(Wrk_AutoAckT.TT) ]OTU(Wrk_Alm);
   // If the Alarm Input (Inp) is true (inverted in EnableInFalse) and the alarm is
   // (or becomes) Enabled, Unsuppressed and Unshelved, this rung sets the Alarm (Alm) bit.
   // The Acknowledge (Ack) bit is cleared when the Alarm initially occurs.
   // #####  V3.0-00  2013-06-30:  Removed Wrk_Abnormal logic.  #####
   // @@@@@  "Inp" is Inverted in the EnableInFalse Routine!  @@@@@
   16: XIO(Inp)XIO(Sts_AlmInh)[XIO(Wrk_Alm) OTU(Ack) ,OTL(Wrk_Alm) ];